HMI tags "Default tag table"
   "buttonView" : Bool, internal
   "messageView" : Bool, internal
   "RPA30R_LCDSwitchAutomat_Manual" : Bool = PLC "RPA30R_LCDSwitchAutomat_Manual", 100 ms
   "RPA30R_light" : Bool = PLC "RPA30R_light", 100 ms
   "RPA30_DataBlock_RPA30_Start" : Bool, 100 ms
   "RPA30_DataBlock_RPA30_scannedFrameBareCode" : String[254], 100 ms
   "RPA30_DataBlock_RPA30_cyclusState" : UInt, 100 ms
   "RPA30_DataBlock_RPA30_scannedData" : String[254], 100 ms
   "outputStatePageChose" : Int, internal
   "ipnut_page_switch" : Int, internal
   "inputStatePageChose" : Int, internal
   "RPA30R_RoofRotationSensorYL" : Bool = PLC "RPA30R_RoofRotationSensorYL", 100 ms
   "RPA30R_RoofRotationSensorYAtOperator" : Bool = PLC "RPA30R_RoofRotationSensorYAtOperator", 100 ms
   "RPA30R_RoofRotationSensorYR" : Bool = PLC "RPA30R_RoofRotationSensorYR", 100 ms
   "RPA30R_RoofRotationSensorYFromOperator" : Bool = PLC "RPA30R_RoofRotationSensorYFromOperator", 100 ms
   "RPA30R_PositionCylinderSensorUnlockY" : Bool = PLC "RPA30R_PositionCylinderSensorUnlockY", 100 ms
   "RPA30R_PositionCylinderSensorLockY" : Bool = PLC "RPA30R_PositionCylinderSensorLockY", 100 ms
   "RPA30R_SensorIFMLeftTriggerOut" : Bool = PLC "RPA30R_SensorIFMLeftTriggerOut", 100 ms
   "RPA30R_SensorIFMLeftReadyOut" : Bool = PLC "RPA30R_SensorIFMLeftReadyOut", 100 ms
   "RPA30R_SensorIFMLeftOut" : Bool = PLC "RPA30R_SensorIFMLeftOut", 100 ms
   "RPA30R_SensorIFMRightTriggerOut" : Bool = PLC "RPA30R_SensorIFMRightTriggerOut", 100 ms
   "RPA30R_SensorIFMRightReadyOut" : Bool = PLC "RPA30R_SensorIFMRightReadyOut", 100 ms
   "RPA30R_SensorIFMRightOut" : Bool = PLC "RPA30R_SensorIFMRightOut", 100 ms
   "RPA30R_ValveCylinderYLock" : Bool = PLC "RPA30R_ValveCylinderYLock", 100 ms
   "RPA30R_SensorIFMLeftTrigger" : Bool = PLC "RPA30R_SensorIFMLeftTrigger", 100 ms
   "RPA30R_SensorIFMLeft_Input_1" : Bool = PLC "RPA30R_SensorIFMLeft_Input_1", 100 ms
   "RPA30R_SensorIFMLeft_Input_2" : Bool = PLC "RPA30R_SensorIFMLeft_Input_2", 100 ms
   "RPA30R_SensorIFMRightTrigger" : Bool = PLC "RPA30R_SensorIFMRightTrigger", 100 ms
   "RPA30R_SensorIFMRight_Input_1" : Bool = PLC "RPA30R_SensorIFMRight_Input_1", 100 ms
   "RPA30R_SensorIFMRight_Input_2" : Bool = PLC "RPA30R_SensorIFMRight_Input_2", 100 ms
   "RPA30R_PrimerPA10SensorPadLeft" : Bool = PLC "RPA30R_PrimerPA10SensorPadLeft", 100 ms
   "RPA30R_PrimerPA10SensorPadRight" : Bool = PLC "RPA30R_PrimerPA10SensorPadRight", 100 ms
   "RPA30R_PrimerPA10SensorFelt" : Bool = PLC "RPA30R_PrimerPA10SensorFelt", 100 ms
   "RPA30R_PrimerPA30SensorRemover208" : Bool = PLC "RPA30R_PrimerPA30SensorRemover208", 100 ms
   "RPA30R_PrimerPA30SensorFeltEmpty" : Bool = PLC "RPA30R_PrimerPA30SensorFeltEmpty", 100 ms
   "RPA30R_LCDButtonStart" : Bool = PLC "RPA30R_LCDButtonStart", 100 ms
   "RPA30R_LCDButtonConfirmSignal" : Bool = PLC "RPA30R_LCDButtonConfirmSignal", 100 ms
   "RPA30R_PrimerPA30SensorBottleRemover208" : Bool = PLC "RPA30R_PrimerPA30SensorBottleRemover208", 100 ms
   "RPA30R_PrimerPA30SensorBottlePrimer207" : Bool = PLC "RPA30R_PrimerPA30SensorBottlePrimer207", 100 ms
   "RPA30R_Beacon_1_LCDPanelGreen" : Bool = PLC "RPA30R_Beacon_1_LCDPanelGreen", 100 ms
   "RPA30R_Beacon_1_LCDPanelOrange" : Bool = PLC "RPA30R_Beacon_1_LCDPanelOrange", 100 ms
   "RPA30R_Beacon_1_LCDPanelRed" : Bool = PLC "RPA30R_Beacon_1_LCDPanelRed", 100 ms
   "RPA30R_Beacon_1_LCDPanelSiren" : Bool = PLC "RPA30R_Beacon_1_LCDPanelSiren", 100 ms
   "RPA30R_Beacon_2_PrimerBoxGreen" : Bool = PLC "RPA30R_Beacon_2_PrimerBoxGreen", 100 ms
   "RPA30R_Beacon_2_PrimerBoxOrange" : Bool = PLC "RPA30R_Beacon_2_PrimerBoxOrange", 100 ms
   "RPA30R_Beacon_2_PrimerBoxRed" : Bool = PLC "RPA30R_Beacon_2_PrimerBoxRed", 100 ms
   "RPA30R_Beacon_2_PrimerBoxSiren" : Bool = PLC "RPA30R_Beacon_2_PrimerBoxSiren", 100 ms
   "RPA30R_PrimerPA30GreenReady" : Bool = PLC "RPA30R_PrimerPA30GreenReady", 100 ms
   "RPA30R_PrimerPA30GreenFelt" : Bool = PLC "RPA30R_PrimerPA30GreenFelt", 100 ms
   "RPA30R_PrimerPA30GreenRemover208" : Bool = PLC "RPA30R_PrimerPA30GreenRemover208", 100 ms
   "RPA30R_PrimerPA30GreenPrimer207" : Bool = PLC "RPA30R_PrimerPA30GreenPrimer207", 100 ms
   "RPA30R_PrimerPA30RedNotReady" : Bool = PLC "RPA30R_PrimerPA30RedNotReady", 100 ms
   "RPA30R_PrimerPA30RedChangePad" : Bool = PLC "RPA30R_PrimerPA30RedChangePad", 100 ms
   "RPA30R_LEDGreenSart" : Bool = PLC "RPA30R_LEDGreenSart", 100 ms
   "RPA30R_LedBlueConfirm" : Bool = PLC "RPA30R_LedBlueConfirm", 100 ms
   "RPA30_DataBlock_RPA30_failStateLock" : Int, 100 ms
   "Clock_0.5Hz" : Bool = PLC "Clock_0.5Hz", 100 ms
   "RPA30_DataBlock_RPA30_bigFailStateLock" : Int, 100 ms
   "RPA30_DataBlock_RPA30_ErrorStateLock" : Int, 100 ms
   "RPA30_DataBlock_RPA30_fatalErrorStateLock" : Int, 100 ms
   "RPA30_IFM_point_checking_DB_points" : Int, 100 ms
   "manual_output_page_switch" : Int, internal
   "input_output_switch" : Bool, internal
   "output_page_switch" : Int, internal
   "PLC_datablock_stations_configuration" : Byte, 1 s
   "configuration_choose" : Int, internal
   "RPA30_DataBlock_RPA30_show_points_hmi" : Byte, 100 ms
   "RPA30_DataBlock_RPA30_actual_instruction_index" : Byte, 1 s
   "RPA30_DataBlock_RPA30_show_smile" : Bool, 100 ms
   "RPA30_DataBlock_RPA30_show_pad_left" : Bool, 100 ms
   "RPA30_DataBlock_RPA30_show_pad_right" : Bool, 100 ms
   "RPA30_DataBlock_pa30_bottle_cyclus_replace" : UInt, 1 s
   "RPA30_DataBlock_pa30_bottle_timing" : LInt, 1 s
   "RPA30_DataBlock_pa30_keyence_switch" : Bool, 1 s

text list "RPA30_InstructionList": 0 ''; 1 ''; 4 ''; 5 ''; 6 ''; 7 ''; 9 ''; 16 ''; 17 ''; 18 ''; 19 ''; 20 ''; 21 ''; 22 ''; 23 ''; 24 ''; 25 ''; 26 ''; 27 ''; 28 ''

text list "pa30_fail_list": 200 ''; 210 ''; 100 ''; 300 ''

text list "PA30_error_list": 1000 ''; 25000 ''; 26000 ''; 24000 ''; 23000 ''; 22000 ''; 400 ''; 401 ''; 402 ''; 403 ''; 155 ''

text list "PA30_fatal_error_list": 150 ''; 160 ''; 190 ''

text list "RPA30_station_configuration": 0 ''; 1 ''; 2 ''

screen "Home" 800x480
   TextField "Text field_3" at 325,5 size 300x40
   TextField "Text field_2" at 2,85 size 70x40
   TextField "Text field_4" at 73,85 size 70x40
   TextField "Text field_5" at 335,130 size 130x25
   TextField "Text field_6" at 20,171 size 330x22
   TextField "Text field_7" at 20,201 size 330x22
   TextField "Text field_8" at 20,231 size 330x22
   TextField "Text field_9" at 20,261 size 330x22
   TextField "Text field_10" at 20,291 size 330x22
   TextField "Text field_11" at 20,321 size 330x22
   TextField "Text field_12" at 20,351 size 330x22
   TextField "Text field_13" at 20,381 size 330x22
   TextField "Text field_14" at 410,171 size 330x22
   TextField "Text field_15" at 410,201 size 330x22
   TextField "Text field_16" at 410,231 size 330x22
   TextField "Text field_17" at 410,261 size 330x22
   TextField "Text field_18" at 410,291 size 330x22
   TextField "Text field_19" at 410,321 size 330x22
   TextField "Text field_20" at 410,351 size 330x22
   TextField "Text field_21" at 410,381 size 330x22
   Button "Button_1" at 640,420 size 80x60
   Button "HmiScreenItemData_1" at 0,420 size 80x60
   Button "HmiScreenItemData_2" at 400,420 size 80x60
   Button "Button_2" at 560,420 size 80x60
   Button "Button_6" at 720,420 size 80x60
   DateTimeField "Date/time field_1" at 650,27 size 150x25
   DateTimeField "Date/time field_2" at 650,0 size 150x28
   TextField "Text field_1" at 0,0 size 300x50
   Button "HmiScreenItemData_3" at 240,420 size 80x60
   Button "HmiScreenItemData_4" at 320,420 size 80x60
   Button "Button_3" at 480,420 size 80x60
   Button "HmiScreenItemData_5" at 80,420 size 80x60
   Button "HmiScreenItemData_6" at 160,420 size 80x60
   Button "Button_11" at 0,420 size 80x60
   Button "Button_12" at 80,420 size 80x60
   Button "Button_13" at 160,420 size 80x60
   Button "Button_14" at 240,420 size 80x60
   Button "Button_15" at 320,420 size 80x60
   Button "Button_16" at 400,420 size 80x60
   Button "Button_17" at 480,420 size 80x60
   Button "Button_18" at 560,420 size 80x60
   Button "Button_19" at 640,420 size 80x60
   Button "Button_20" at 720,420 size 80x60
   TextField "Text field_22" at 64,67 size 129x22
   AlarmView "Alarm view_1" at 60,90 size 680x320
   Button "Button_9" at 715,65 size 25x25
   TextField "Text field_37" at 360,54 size 120x25

screen "I0-State" 800x480
   TextField "Text field_3" at 325,5 size 300x40
   Button "Button_1" at 640,420 size 80x60
   Button "Button_4" at 160,420 size 80x60
   Button "HmiScreenItemData_3" at 400,420 size 80x60
   Button "Button_2" at 560,420 size 80x60
   Button "Button_6" at 720,420 size 80x60
   Button "HmiScreenItemData_2" at 240,420 size 80x60
   Button "HmiScreenItemData_4" at 320,420 size 80x60
   TextField "Text field_1" at 0,0 size 300x50
   DateTimeField "Date/time field_2" at 650,0 size 150x28
   DateTimeField "Date/time field_1" at 650,27 size 150x25
   Button "HmiScreenItemData_1" at 0,420 size 80x60
   Button "Button_3" at 480,420 size 80x60
   Button "Button_5" at 80,420 size 80x60
   Button "input_back" at 20,52 size 90x25
   Button "input_next" at 690,52 size 90x25
   Button "output_back" at 20,52 size 90x25
   Button "output_next" at 690,52 size 90x25
   TextField "Text field_2" at 20,85 size 330x22
   TextField "Text field_4" at 20,115 size 330x22
   TextField "Text field_5" at 20,145 size 330x22
   TextField "Text field_6" at 20,175 size 330x22
   TextField "Text field_7" at 20,205 size 330x22
   TextField "Text field_8" at 20,235 size 330x22
   TextField "Text field_9" at 20,265 size 330x22
   TextField "Text field_10" at 20,295 size 330x22
   TextField "Text field_11" at 20,325 size 330x22
   TextField "Text field_12" at 20,355 size 330x22
   TextField "Text field_13" at 20,385 size 330x22
   TextField "Text field_14" at 410,85 size 330x22
   TextField "Text field_15" at 410,115 size 330x22
   TextField "Text field_16" at 410,145 size 330x22
   TextField "Text field_17" at 410,175 size 330x22
   TextField "Text field_18" at 410,205 size 330x22
   TextField "Text field_19" at 410,235 size 330x22
   TextField "Text field_20" at 410,265 size 330x22
   TextField "Text field_21" at 410,295 size 330x22
   TextField "Text field_22" at 410,325 size 330x22
   TextField "Text field_23" at 410,355 size 330x22
   TextField "Text field_24" at 410,385 size 330x22
   Button "Button_11" at 0,420 size 80x60
   Button "Button_12" at 80,420 size 80x60
   Button "Button_13" at 160,420 size 80x60
   Button "Button_14" at 240,420 size 80x60
   Button "Button_15" at 320,420 size 80x60
   Button "Button_16" at 400,420 size 80x60
   Button "Button_17" at 480,420 size 80x60
   Button "Button_18" at 560,420 size 80x60
   Button "Button_19" at 640,420 size 80x60
   Button "Button_20" at 720,420 size 80x60
   TextField "Text field_25" at 64,67 size 129x22
   AlarmView "Alarm view_1" at 60,90 size 680x320
   Button "Button_9" at 715,65 size 25x25
   TextField "Text field_26" at 20,85 size 330x22
   TextField "Text field_27" at 20,115 size 330x22
   TextField "Text field_28" at 20,145 size 330x22
   TextField "Text field_29" at 20,175 size 330x22
   TextField "Text field_30" at 20,205 size 330x22
   TextField "Text field_31" at 20,235 size 330x22
   TextField "Text field_32" at 20,265 size 330x22
   TextField "Text field_33" at 20,295 size 330x22
   TextField "Text field_34" at 20,325 size 330x22
   TextField "Text field_35" at 20,355 size 330x22
   TextField "Text field_36" at 20,385 size 330x22
   TextField "Text field_37" at 410,85 size 330x22
   TextField "Text field_38" at 410,115 size 330x22
   TextField "Text field_39" at 410,145 size 330x22
   TextField "Text field_40" at 410,175 size 330x22
   TextField "Text field_41" at 410,205 size 330x22
   TextField "Text field_42" at 410,235 size 330x22
   TextField "Text field_43" at 410,265 size 330x22
   TextField "Text field_44" at 410,295 size 330x22
   TextField "Text field_45" at 410,325 size 330x22
   TextField "Text field_46" at 410,355 size 330x22
   TextField "Text field_47" at 410,385 size 330x22
   TextField "Text field_48" at 20,85 size 330x22
   TextField "Text field_49" at 20,85 size 330x22
   TextField "Text field_50" at 360,54 size 120x25

screen "Main_page" 800x480
   Button "HmiScreenItemData_1" at 80,420 size 80x60
   TextField "Text field_2" at 0,85 size 800x25
   TextField "Text field_3" at 325,5 size 300x40
   Button "Button_4" at 480,420 size 80x60
   Button "Button_5" at 640,420 size 80x60
   Button "Button_1" at 0,420 size 80x60
   Button "Button_7" at 400,420 size 80x60
   Button "HmiScreenItemData_2" at 160,420 size 80x60
   Button "Button_3" at 560,420 size 80x60
   Button "Button_6" at 720,420 size 80x60
   Button "HmiScreenItemData_3" at 240,420 size 80x60
   Button "HmiScreenItemData_4" at 320,420 size 80x60
   TextField "Text field_1" at 0,0 size 300x50
   DateTimeField "Date/time field_2" at 650,0 size 150x28
   DateTimeField "Date/time field_1" at 650,27 size 150x25
   SymbolicIOField "Symbolic I/O field_1" at 10,110 size 780x90
   Button "HmiScreenItemData_5" at 80,420 size 80x60
   SymbolicIOField "Symbolic I/O field_6" at 171,50 size 169x32
   TextField "Text field_56" at 11,51 size 143x27
   Button "Button_2" at 400,420 size 80x60
   Button "Button_11" at 0,420 size 80x60
   Button "Button_12" at 80,420 size 80x60
   Button "Button_13" at 160,420 size 80x60
   Button "Button_14" at 240,420 size 80x60
   Button "Button_15" at 320,420 size 80x60
   Button "Button_16" at 400,420 size 80x60
   Button "Button_17" at 480,420 size 80x60
   Button "Button_18" at 560,420 size 80x60
   Button "Button_19" at 640,420 size 80x60
   Button "Button_20" at 720,420 size 80x60
   GraphicView "Graphic view_1" at 320,228 size 180x180
   TextField "Text field_5" at 64,67 size 129x22
   AlarmView "Alarm view_1" at 60,90 size 680x320
   Button "Button_9" at 715,65 size 25x25
   SymbolicIOField "Symbolic I/O field_2" at 0,170 size 800x110
   SymbolicIOField "Symbolic I/O field_3" at 0,170 size 800x110
   SymbolicIOField "Symbolic I/O field_4" at 0,170 size 800x110
   SymbolicIOField "Symbolic I/O field_5" at 0,170 size 800x110
   TextField "Text field_10" at 165,322 size 22x37
   TextField "Text field_11" at 279,323 size 22x37
   TextField "Text field_12" at 392,323 size 22x37
   TextField "Text field_13" at 494,322 size 22x37
   TextField "Text field_14" at 613,323 size 22x37
   TextField "Text field_6" at 163,255 size 22x37
   TextField "Text field_7" at 392,255 size 22x37
   TextField "Text field_8" at 613,255 size 22x37
   TextField "Text field_37" at 360,54 size 120x25
   GraphicView "Graphic view_2" at 207,225 size 345x187
   GraphicView "Graphic view_3" at 260,225 size 345x187
   TextField "Text field_4" at 299,290 size 237x43

screen "Scanner" 800x480
   TextField "Text field_3" at 325,5 size 300x40
   IOField "I/O field_1" at 10,118 size 780x32
   TextField "Text field_2" at 10,86 size 141x22
   Button "Button_1" at 640,420 size 80x60
   Button "HmiScreenItemData_3" at 400,420 size 80x60
   Button "Button_2" at 560,420 size 80x60
   Button "Button_6" at 720,420 size 80x60
   DateTimeField "Date/time field_2" at 650,0 size 150x28
   TextField "Text field_1" at 0,0 size 300x50
   DateTimeField "Date/time field_1" at 650,27 size 150x25
   Button "HmiScreenItemData_2" at 240,420 size 80x60
   Button "HmiScreenItemData_4" at 320,420 size 80x60
   Button "HmiScreenItemData_1" at 0,420 size 80x60
   Button "HmiScreenItemData_5" at 480,420 size 80x60
   Button "HmiScreenItemData_6" at 160,420 size 80x60
   Button "HmiScreenItemData_7" at 80,420 size 80x60
   Button "Button_3" at 27,167 size 96x32
   Button "Button_11" at 0,420 size 80x60
   Button "Button_12" at 80,420 size 80x60
   Button "Button_13" at 160,420 size 80x60
   Button "Button_14" at 240,420 size 80x60
   Button "Button_15" at 320,420 size 80x60
   Button "Button_16" at 400,420 size 80x60
   Button "Button_17" at 480,420 size 80x60
   Button "Button_18" at 560,420 size 80x60
   Button "Button_19" at 640,420 size 80x60
   Button "Button_20" at 720,420 size 80x60
   TextField "Text field_5" at 64,67 size 129x22
   AlarmView "Alarm view_1" at 60,90 size 680x320
   Button "Button_9" at 715,65 size 25x25
   TextField "Text field_37" at 360,54 size 120x25

screen "Manual" 800x480
   TextField "Text field_3" at 325,5 size 300x40
   Button "Button_4" at 18,85 size 50x50
   Button "Button_12" at 730,85 size 50x50
   Button "Button_1" at 640,420 size 80x60
   Button "HmiScreenItemData_1" at 0,420 size 80x60
   Button "Button_6" at 720,420 size 80x60
   Button "Button_34" at 400,420 size 80x60
   Button "HmiScreenItemData_3" at 240,420 size 80x60
   Button "HmiScreenItemData_4" at 320,420 size 80x60
   TextField "Text field_1" at 0,0 size 300x50
   DateTimeField "Date/time field_2" at 650,0 size 150x28
   DateTimeField "Date/time field_1" at 650,27 size 150x25
   Button "Button_5" at 160,420 size 80x60
   Button "Button_3" at 480,420 size 80x60
   Button "Button_7" at 80,420 size 80x60
   Button "Button_2" at 560,420 size 80x60
   Button "Button_23" at 0,420 size 80x60
   Button "Button_24" at 80,420 size 80x60
   Button "Button_25" at 160,420 size 80x60
   Button "Button_26" at 240,420 size 80x60
   Button "Button_27" at 320,420 size 80x60
   Button "Button_28" at 400,420 size 80x60
   Button "Button_29" at 480,420 size 80x60
   Button "Button_30" at 560,420 size 80x60
   Button "Button_31" at 640,420 size 80x60
   Button "Button_32" at 720,420 size 80x60
   TextField "Text field_8" at 64,67 size 129x22
   AlarmView "Alarm view_1" at 60,90 size 680x320
   Button "Button_33" at 715,65 size 25x25
   Switch "Switch_15" at 717,149 size 64x32
   Switch "Switch_16" at 717,185 size 64x32
   Switch "Switch_17" at 717,221 size 64x32
   Switch "Switch_18" at 717,257 size 64x32
   Switch "Switch_19" at 717,293 size 64x32
   Switch "Switch_20" at 718,328 size 64x32
   Switch "Switch_21" at 719,364 size 64x32
   TextField "Text field_22" at 493,149 size 200x32
   TextField "Text field_23" at 493,181 size 200x32
   TextField "Text field_24" at 492,221 size 200x32
   TextField "Text field_25" at 493,289 size 200x32
   TextField "Text field_26" at 493,257 size 200x32
   TextField "Text field_27" at 493,328 size 200x32
   TextField "Text field_28" at 493,360 size 200x32
   Switch "Switch_22" at 300,149 size 64x32
   Switch "Switch_23" at 300,185 size 64x32
   Switch "Switch_24" at 300,221 size 64x32
   Switch "Switch_25" at 300,257 size 64x32
   Switch "Switch_26" at 300,293 size 64x32
   Switch "Switch_27" at 301,328 size 64x32
   Switch "Switch_28" at 302,364 size 64x32
   TextField "Text field_29" at 76,149 size 200x32
   TextField "Text field_30" at 76,181 size 200x32
   TextField "Text field_31" at 75,221 size 200x32
   TextField "Text field_32" at 76,289 size 200x32
   TextField "Text field_33" at 76,257 size 200x32
   TextField "Text field_34" at 76,328 size 200x32
   TextField "Text field_35" at 76,360 size 200x32
   Switch "Switch_1" at 717,149 size 64x32
   Switch "Switch_2" at 717,185 size 64x32
   TextField "Text field_7" at 493,149 size 200x32
   TextField "Text field_9" at 493,181 size 200x32
   Switch "Switch_8" at 300,149 size 64x32
   Switch "Switch_9" at 300,185 size 64x32
   Switch "Switch_10" at 300,221 size 64x32
   Switch "Switch_11" at 300,257 size 64x32
   Switch "Switch_12" at 300,293 size 64x32
   Switch "Switch_13" at 301,328 size 64x32
   Switch "Switch_14" at 302,364 size 64x32
   TextField "Text field_15" at 76,149 size 200x32
   TextField "Text field_16" at 76,181 size 200x32
   TextField "Text field_17" at 75,221 size 200x32
   TextField "Text field_18" at 37,289 size 239x32
   TextField "Text field_19" at 26,257 size 250x32
   TextField "Text field_20" at 29,328 size 247x32
   TextField "Text field_21" at 44,360 size 232x32
   TextField "Text field_37" at 360,54 size 120x25

screen "System" 800x480
   TextField "Text field_3" at 325,5 size 300x40
   TextField "Text field_2" at 300,86 size 200x27
   Button "Button_4" at 10,290 size 170x60
   Button "Button_5" at 10,355 size 170x60
   Button "Button_7" at 213,290 size 170x60
   Button "Button_8" at 416,290 size 170x60
   Button "Button_9" at 620,290 size 170x60
   Button "Button_11" at 213,355 size 170x60
   Button "Button_12" at 416,355 size 170x60
   Button "Button_13" at 620,355 size 170x60
   AlarmView "Alarm view_1" at 10,115 size 780x170
   Button "HmiScreenItemData_1" at 0,420 size 80x60
   Button "Button_3" at 160,420 size 80x60
   Button "Button_14" at 240,420 size 80x60
   Button "Button_15" at 320,420 size 80x60
   Button "Button_16" at 400,420 size 80x60
   Button "Button_2" at 560,420 size 80x60
   Button "Button_1" at 640,420 size 80x60
   Button "Button_6" at 720,420 size 80x60
   TextField "Text field_1" at 0,0 size 300x50
   DateTimeField "Date/time field_2" at 650,0 size 150x28
   DateTimeField "Date/time field_1" at 650,27 size 150x25
   Button "Button_10" at 80,420 size 80x60
   Button "Button_17" at 480,420 size 80x60
   TextField "Text field_37" at 360,54 size 120x25

screen "Station_configuration" 800x480
   TextField "Text field_3" at 325,5 size 300x40
   Button "Button_1" at 640,420 size 80x60
   Button "HmiScreenItemData_1" at 0,420 size 80x60
   Button "Button_6" at 720,420 size 80x60
   Button "Button_34" at 400,420 size 80x60
   Button "HmiScreenItemData_4" at 320,420 size 80x60
   TextField "Text field_1" at 0,0 size 300x50
   DateTimeField "Date/time field_2" at 650,0 size 150x28
   DateTimeField "Date/time field_1" at 650,27 size 150x25
   Button "Button_5" at 160,420 size 80x60
   Button "Button_3" at 480,420 size 80x60
   Button "Button_7" at 80,420 size 80x60
   Button "Button_2" at 560,420 size 80x60
   SymbolicIOField "Symbolic I/O field_1" at 33,194 size 310x65
   TextField "Text field_2" at 33,159 size 192x27
   Button "Button_4" at 355,195 size 90x65
   SymbolicIOField "Symbolic I/O field_2" at 457,195 size 310x65
   TextField "Text field_4" at 457,159 size 225x27
   Switch "Switch_1" at 370,326 size 64x32
   TextField "Text field_5" at 222,288 size 223x23
   Button "HmiScreenItemData_2" at 240,420 size 80x60
   TextField "Text field_37" at 360,54 size 120x25

screen "chemical_setup" 800x480
   Button "HmiScreenItemData_3" at 400,420 size 80x60
   Button "Button_2" at 560,420 size 80x60
   Button "Button_6" at 720,420 size 80x60
   DateTimeField "Date/time field_2" at 650,0 size 150x28
   TextField "Text field_1" at 0,0 size 300x50
   DateTimeField "Date/time field_1" at 650,27 size 150x25
   Button "HmiScreenItemData_2" at 240,420 size 80x60
   Button "HmiScreenItemData_4" at 320,420 size 80x60
   Button "HmiScreenItemData_1" at 0,420 size 80x60
   Button "HmiScreenItemData_5" at 480,420 size 80x60
   Button "HmiScreenItemData_6" at 160,420 size 80x60
   Button "HmiScreenItemData_7" at 80,420 size 80x60
   IOField "I/O field_1" at 87,130 size 341x44
   IOField "I/O field_2" at 87,237 size 338x44
   TextField "Text field_2" at 85,100 size 137x25
   TextField "Text field_3" at 87,206 size 111x25
   TextField "Text field_4" at 435,245 size 93x20
   Button "Button_1" at 640,420 size 80x60
   Button "Button_11" at 0,420 size 80x60
   Button "Button_12" at 80,420 size 80x60
   Button "Button_13" at 160,420 size 80x60
   Button "Button_14" at 240,420 size 80x60
   Button "Button_15" at 320,420 size 80x60
   Button "Button_16" at 400,420 size 80x60
   Button "Button_17" at 480,420 size 80x60
   Button "Button_18" at 560,420 size 80x60
   Button "Button_19" at 640,420 size 80x60
   Button "Button_20" at 720,420 size 80x60
   TextField "Text field_5" at 64,67 size 129x22
   Button "Button_9" at 715,65 size 25x25
   AlarmView "Alarm view_1" at 60,90 size 680x320
   TextField "Text field_37" at 360,54 size 120x25

screen "User_management" 800x480
   TextField "Text field_3" at 325,5 size 300x40
   Button "HmiScreenItemData_1" at 0,420 size 80x60
   Button "Button_3" at 160,420 size 80x60
   Button "Button_14" at 240,420 size 80x60
   Button "Button_15" at 320,420 size 80x60
   Button "Button_16" at 400,420 size 80x60
   Button "Button_17" at 480,420 size 80x60
   Button "Button_2" at 560,420 size 80x60
   Button "Button_1" at 640,420 size 80x60
   TextField "Text field_1" at 0,0 size 300x50
   DateTimeField "Date/time field_2" at 650,0 size 150x28
   DateTimeField "Date/time field_1" at 650,27 size 150x25
   Button "Button_10" at 80,420 size 80x60
   UserView "User view_1" at 20,92 size 758x304
   Button "Button_4" at 720,420 size 80x60
   TextField "Text field_37" at 360,54 size 120x25
*)

(* ===== HMI "HMI_RT_4" =====
connection "HMI_Connection_4": ETHERNET, SMART_S7_1500_OMS

HMI tags "Default tag table"
   "buttonView" : Bool, internal
   "messageView" : Bool, internal
   "RPA60R_LCDSwitchAutomat_Manual" : Bool = PLC "RPA60R_LCDSwitchAutomat_Manual", 100 ms
   "RPA60R_light" : Bool = PLC "RPA60R_light", 100 ms
   "RPA60_DataBlock_RPA60_Start" : Bool, 100 ms
   "RPA60_DataBlock_RPA60_cyclusState" : UInt, 100 ms
   "RPA60_DataBlock_RPA60_scannedFrameBareCode" : String[254], 100 ms
   "RPA60_DataBlock_RPA60_failStateLock" : Int, 100 ms
   "RPA60_DataBlock_RPA60_scanedData" : String[254], 100 ms
   "inputOutputStatePageChose" : Int, internal
   "RPA60R_RoofRotationSensorYL" : Bool = PLC "RPA60R_RoofRotationSensorYL", 100 ms
   "RPA60R_RoofRotationSensorYAtOperator" : Bool = PLC "RPA60R_RoofRotationSensorYAtOperator", 100 ms
   "RPA60R_RoofRotationSensorYR" : Bool = PLC "RPA60R_RoofRotationSensorYR", 100 ms
   "RPA60R_RoofRotationSensorYFromOperator" : Bool = PLC "RPA60R_RoofRotationSensorYFromOperator", 100 ms
   "RPA60R_valvePositionSensorUnlockY" : Bool = PLC "RPA60R_valvePositionSensorUnlockY", 100 ms
   "RPA60R_valvePositionSensorLockY" : Bool = PLC "RPA60R_valvePositionSensorLockY", 100 ms
   "RPA60R_SenzorLoaderPresenceLeft581" : Bool = PLC "RPA60R_SenzorLoaderPresenceLeft581", 100 ms
   "RPA60R_SenzorLoaderPresenceRight581" : Bool = PLC "RPA60R_SenzorLoaderPresenceRight581", 100 ms
   "RPA60R_SenzorLoaderPresenceLeft582" : Bool = PLC "RPA60R_SenzorLoaderPresenceLeft582", 100 ms
   "RPA60R_SenzorLoaderPresenceRear582" : Bool = PLC "RPA60R_SenzorLoaderPresenceRear582", 100 ms
   "RPA60R_SenzorLoaderPresenceRight582" : Bool = PLC "RPA60R_SenzorLoaderPresenceRight582", 100 ms
   "RPA60R_SenzorSealPresenceLeft581" : Bool = PLC "RPA60R_SenzorSealPresenceLeft581", 100 ms
   "RPA60R_SenzorSealPresenceRear581" : Bool = PLC "RPA60R_SenzorSealPresenceRear581", 100 ms
   "RPA60R_SenzorSealPresenceRight581" : Bool = PLC "RPA60R_SenzorSealPresenceRight581", 100 ms
   "RPA60R_SenzorSealPresenceLeft582" : Bool = PLC "RPA60R_SenzorSealPresenceLeft582", 100 ms
   "RPA60R_SenzorSealPresenceRear582" : Bool = PLC "RPA60R_SenzorSealPresenceRear582", 100 ms
   "RPA60R_SenzorSealPresenceRight582" : Bool = PLC "RPA60R_SenzorSealPresenceRight582", 100 ms
   "RPA60R_SenzorVacuum" : Bool = PLC "RPA60R_SenzorVacuum", 100 ms
   "RPA60R_ValveCylinderYLock" : Bool = PLC "RPA60R_ValveCylinderYLock", 100 ms
   "RPA60R_LCDButtonStart" : Bool = PLC "RPA60R_LCDButtonStart", 100 ms
   "RPA60R_LCDButtonConfirmSignal" : Bool = PLC "RPA60R_LCDButtonConfirmSignal", 100 ms
   "RPA60R_Beacon_1_LCDPanelGreen" : Bool = PLC "RPA60R_Beacon_1_LCDPanelGreen", 100 ms
   "RPA60R_Beacon_1_LCDPanelOrange" : Bool = PLC "RPA60R_Beacon_1_LCDPanelOrange", 100 ms
   "RPA60R_Beacon_1_LCDPanelRed" : Bool = PLC "RPA60R_Beacon_1_LCDPanelRed", 100 ms
   "RPA60R_Beacon_1_LCDPanelSiren" : Bool = PLC "RPA60R_Beacon_1_LCDPanelSiren", 100 ms
   "RPA60R_LEDGreenSart" : Bool = PLC "RPA60R_LEDGreenSart", 100 ms
   "RPA60R_LedBlueConfirm" : Bool = PLC "RPA60R_LedBlueConfirm", 100 ms
   "RPA60R_VacuumSwitch" : Bool = PLC "RPA60R_VacuumSwitch", 100 ms
   "RPA60R_LEDRoller" : Bool = PLC "RPA60R_LEDRoller", 100 ms
   "RPA60R_SenzorRoller" : Bool = PLC "RPA60R_SenzorRoller", 100 ms
   "RPA30R_Beacon_1_LCDPanelSiren" : Bool = PLC "RPA30R_Beacon_1_LCDPanelSiren", 100 ms
   "RPA60_DataBlock_RPA60_bigFailStateLock" : Int, 1 s
   "RPA60_DataBlock_RPA60_fatalErrorStateLock" : Int, 1 s
   "RPA60_DataBlock_RPA60_ErrorStateLock" : Int, 1 s
   "Clock_0.5Hz" : Bool = PLC "Clock_0.5Hz", 1 s
   "RPA60_DataBlock_RPA60_printEnable" : Bool, 1 s
   "input_output_switch" : Bool, internal
   "output_switch_page" : Int, internal
   "input_switch_page" : Int, internal
   "PLC_datablock_stations_configuration" : Byte, 1 s
   "RPA60_DataBlock_RPA60_hmi_instruction_index" : Byte, 1 s
   "RPA60_DataBlock_RPA60_show_smile" : Bool, 1 s
   "RPA60_DataBlock_RPA60_number_of_check" : Byte, 1 s
   "RPA60_DataBlock_RPA60_show_check_button" : Bool, 1 s
   "RPA60_DataBlock_RPA60_station_configuration" : Byte, 1 s
   "choose_configuration" : Int, internal
   "RPA60_DataBlock_RPA60_hardware_configuration" : Byte, 1 s
   "DB_RPA60_CAM_RPA60_ENABLE_CAMERAS" : Bool, 500 ms

text list "PA60_instructionList": 0 ''; 3 ''; 7 ''; 8 ''; 9 ''; 24 ''; 26 ''; 27 ''; 23 ''; 28 ''; 11 ''; 29 ''; 30 ''; 39 ''; 40 ''; 41 ''

text list "PA60_error_list": 1000 ''; 26000 ''; 25000 ''; 24000 ''; 23000 ''; 20000 ''; 21000 ''; 27000 ''

text list "PA60_fatal_error_list": 170 ''; 150 ''; 180 ''; 230 ''; 293 ''; 294 ''; 190 ''

text list "PA60_big_fail_list": 120 ''

text list "RPA60_station_configuration": 0 ''; 1 ''; 2 ''

text list "RPA60_hardware_configuration": 0 ''; 1 ''; 3..255 ''; 2 ''

screen "Home" 800x480
   TextField "Text field_3" at 325,5 size 300x40
   TextField "Text field_2" at 2,85 size 70x40
   TextField "Text field_5" at 335,130 size 130x25
   TextField "Text field_6" at 20,171 size 330x22
   TextField "Text field_7" at 20,201 size 330x22
   Button "Button_1" at 640,420 size 80x60
   Button "HmiScreenItemData_1" at 0,420 size 80x60
   Button "HmiScreenItemData_2" at 400,420 size 80x60
   Button "Button_2" at 560,420 size 80x60
   Button "Button_6" at 720,420 size 80x60
   DateTimeField "Date/time field_1" at 650,27 size 150x25
   DateTimeField "Date/time field_2" at 650,0 size 150x28
   TextField "Text field_1" at 0,0 size 300x50
   Button "HmiScreenItemData_3" at 240,420 size 80x60
   Button "HmiScreenItemData_4" at 320,420 size 80x60
   Button "Button_3" at 480,420 size 80x60
   Button "HmiScreenItemData_5" at 80,420 size 80x60
   Button "HmiScreenItemData_6" at 160,420 size 80x60
   IOField "I/O field_1" at 73,85 size 70x40
   Button "Button_11" at 0,420 size 80x60
   Button "Button_12" at 80,420 size 80x60
   Button "Button_13" at 160,420 size 80x60
   Button "Button_14" at 240,420 size 80x60
   Button "Button_15" at 320,420 size 80x60
   Button "Button_16" at 400,420 size 80x60
   Button "Button_17" at 480,420 size 80x60
   Button "Button_18" at 560,420 size 80x60
   Button "Button_19" at 640,420 size 80x60
   Button "Button_20" at 720,420 size 80x60
   TextField "Text field_22" at 64,67 size 129x22
   AlarmView "Alarm view_1" at 60,90 size 680x320
   Button "Button_9" at 715,65 size 25x25
   TextField "Text field_37" at 360,54 size 120x25

screen "I0-State" 800x480
   TextField "Text field_3" at 325,5 size 300x40
   Button "Button_1" at 640,420 size 80x60
   Button "Button_4" at 160,420 size 80x60
   Button "HmiScreenItemData_3" at 400,420 size 80x60
   Button "Button_2" at 560,420 size 80x60
   Button "Button_6" at 720,420 size 80x60
   Button "HmiScreenItemData_2" at 240,420 size 80x60
   Button "HmiScreenItemData_4" at 320,420 size 80x60
   TextField "Text field_1" at 0,0 size 300x50
   DateTimeField "Date/time field_2" at 650,0 size 150x28
   DateTimeField "Date/time field_1" at 650,27 size 150x25
   Button "HmiScreenItemData_1" at 0,420 size 80x60
   Button "Button_3" at 480,420 size 80x60
   Button "Button_5" at 80,420 size 80x60
   Button "input_back" at 20,52 size 90x25
   Button "input_next" at 690,52 size 90x25
   Button "output_back" at 20,52 size 90x25
   Button "output_next" at 690,52 size 90x25
   TextField "Text field_2" at 20,85 size 330x22
   TextField "Text field_4" at 20,115 size 330x22
   TextField "Text field_5" at 20,145 size 330x22
   TextField "Text field_6" at 20,175 size 330x22
   TextField "Text field_7" at 20,205 size 330x22
   TextField "Text field_8" at 20,235 size 330x22
   TextField "Text field_9" at 20,265 size 330x22
   TextField "Text field_10" at 20,295 size 330x22
   TextField "Text field_11" at 20,325 size 330x22
   TextField "Text field_12" at 20,355 size 330x22
   TextField "Text field_13" at 20,385 size 330x22
   TextField "Text field_14" at 410,85 size 330x22
   TextField "Text field_15" at 410,115 size 330x22
   TextField "Text field_16" at 410,145 size 330x22
   TextField "Text field_17" at 410,175 size 330x22
   TextField "Text field_18" at 410,205 size 330x22
   TextField "Text field_19" at 410,235 size 330x22
   TextField "Text field_20" at 410,265 size 330x22
   TextField "Text field_21" at 410,295 size 330x22
   TextField "Text field_22" at 410,325 size 330x22
   TextField "Text field_23" at 410,355 size 330x22
   TextField "Text field_24" at 410,385 size 330x22
   Button "Button_11" at 0,420 size 80x60
   Button "Button_12" at 80,420 size 80x60
   Button "Button_13" at 160,420 size 80x60
   Button "Button_14" at 240,420 size 80x60
   Button "Button_15" at 320,420 size 80x60
   Button "Button_16" at 400,420 size 80x60
   Button "Button_17" at 480,420 size 80x60
   Button "Button_18" at 560,420 size 80x60
   Button "Button_19" at 640,420 size 80x60
   Button "Button_20" at 720,420 size 80x60
   TextField "Text field_25" at 64,67 size 129x22
   AlarmView "Alarm view_1" at 60,90 size 680x320
   Button "Button_9" at 715,65 size 25x25
   TextField "Text field_26" at 20,85 size 330x22
   TextField "Text field_27" at 20,115 size 330x22
   TextField "Text field_28" at 20,145 size 330x22
   TextField "Text field_29" at 20,175 size 330x22
   TextField "Text field_30" at 20,205 size 330x22
   TextField "Text field_31" at 20,235 size 330x22
   TextField "Text field_32" at 20,265 size 330x22
   TextField "Text field_33" at 20,295 size 330x22
   TextField "Text field_34" at 20,325 size 330x22
   TextField "Text field_48" at 21,85 size 330x22
   TextField "Text field_37" at 360,54 size 120x25

screen "Main_page" 800x480
   Button "HmiScreenItemData_1" at 80,420 size 80x60
   TextField "Text field_2" at 0,85 size 800x25
   TextField "Text field_3" at 325,5 size 300x40
   Button "Button_4" at 480,420 size 80x60
   Button "Button_5" at 640,420 size 80x60
   Button "Button_1" at 0,420 size 80x60
   Button "HmiScreenItemData_2" at 160,420 size 80x60
   Button "Button_2" at 400,420 size 80x60
   Button "Button_3" at 560,420 size 80x60
   Button "Button_6" at 720,420 size 80x60
   Button "HmiScreenItemData_3" at 240,420 size 80x60
   Button "HmiScreenItemData_4" at 320,420 size 80x60
   TextField "Text field_1" at 0,0 size 300x50
   DateTimeField "Date/time field_2" at 650,0 size 150x28
   DateTimeField "Date/time field_1" at 650,27 size 150x25
   SymbolicIOField "Symbolic I/O field_1" at 10,110 size 780x90
   Button "HmiScreenItemData_5" at 80,420 size 80x60
   GraphicView "Graphic view_1" at 320,228 size 180x180
   SymbolicIOField "Symbolic I/O field_6" at 169,51 size 169x32
   TextField "Text field_56" at 12,52 size 143x27
   Button "Button_21" at 720,420 size 80x60
   Button "Button_22" at 400,420 size 80x60
   Button "Button_11" at 0,420 size 80x60
   Button "Button_13" at 160,420 size 80x60
   Button "Button_14" at 240,420 size 80x60
   Button "Button_15" at 320,420 size 80x60
   Button "Button_16" at 400,420 size 80x60
   Button "Button_17" at 480,420 size 80x60
   Button "Button_18" at 560,420 size 80x60
   Button "Button_19" at 640,420 size 80x60
   Button "Button_20" at 720,420 size 80x60
   Button "Button_12" at 80,420 size 80x60
   TextField "Text field_5" at 64,67 size 129x22
   AlarmView "Alarm view_1" at 60,90 size 680x320
   Button "Button_9" at 715,65 size 25x25
   SymbolicIOField "Symbolic I/O field_2" at 0,170 size 800x110
   SymbolicIOField "Symbolic I/O field_3" at 0,170 size 800x110
   SymbolicIOField "Symbolic I/O field_4" at 0,170 size 800x110
   SymbolicIOField "Symbolic I/O field_5" at 0,170 size 800x110
   Button "Button_7" at 486,333 size 130x50
   Button "Button_10" at 213,333 size 130x50
   Button "Button_8" at 350,333 size 130x50
   TextField "Text field_37" at 360,54 size 120x25
   TextField "Text field_4" at 302,290 size 237x43

screen "Scanner" 800x480
   TextField "Text field_3" at 325,5 size 300x40
   IOField "I/O field_1" at 10,120 size 780x32
   TextField "Text field_2" at 10,88 size 141x22
   Button "Button_1" at 640,420 size 80x60
   Button "HmiScreenItemData_3" at 400,420 size 80x60
   Button "Button_2" at 560,420 size 80x60
   Button "Button_6" at 720,420 size 80x60
   DateTimeField "Date/time field_2" at 650,0 size 150x28
   TextField "Text field_1" at 0,0 size 300x50
   DateTimeField "Date/time field_1" at 650,27 size 150x25
   Button "HmiScreenItemData_2" at 240,420 size 80x60
   Button "HmiScreenItemData_4" at 320,420 size 80x60
   Button "HmiScreenItemData_1" at 0,420 size 80x60
   Button "HmiScreenItemData_5" at 480,420 size 80x60
   Button "HmiScreenItemData_6" at 160,420 size 80x60
   Button "HmiScreenItemData_7" at 80,420 size 80x60
   Button "Button_3" at 10,165 size 96x32
   Button "Button_11" at 0,420 size 80x60
   Button "Button_12" at 80,420 size 80x60
   Button "Button_13" at 160,420 size 80x60
   Button "Button_14" at 240,420 size 80x60
   Button "Button_15" at 320,420 size 80x60
   Button "Button_16" at 400,420 size 80x60
   Button "Button_17" at 480,420 size 80x60
   Button "Button_18" at 560,420 size 80x60
   Button "Button_19" at 640,420 size 80x60
   Button "Button_20" at 720,420 size 80x60
   TextField "Text field_5" at 64,67 size 129x22
   AlarmView "Alarm view_1" at 60,90 size 680x320
   Button "Button_9" at 715,65 size 25x25
   TextField "Text field_37" at 360,54 size 120x25

screen "Manual" 800x480
   TextField "Text field_3" at 325,5 size 300x40
   Button "Button_12" at 730,85 size 50x50
   Button "Button_1" at 640,420 size 80x60
   Button "HmiScreenItemData_1" at 0,420 size 80x60
   Button "Button_2" at 560,420 size 80x60
   Button "Button_6" at 720,420 size 80x60
   Button "Button_34" at 400,420 size 80x60
   Button "HmiScreenItemData_3" at 240,420 size 80x60
   Button "HmiScreenItemData_4" at 320,420 size 80x60
   DateTimeField "Date/time field_2" at 650,0 size 150x28
   DateTimeField "Date/time field_1" at 650,27 size 150x25
   Button "Button_5" at 160,420 size 80x60
   Button "Button_3" at 480,420 size 80x60
   Button "Button_7" at 80,420 size 80x60
   Button "Button_4" at 21,85 size 50x50
   TextField "Text field_1" at 0,0 size 300x50
   Button "Button_23" at 0,420 size 80x60
   Button "Button_24" at 80,420 size 80x60
   Button "Button_25" at 160,420 size 80x60
   Button "Button_26" at 240,420 size 80x60
   Button "Button_27" at 320,420 size 80x60
   Button "Button_28" at 400,420 size 80x60
   Button "Button_29" at 480,420 size 80x60
   Button "Button_30" at 560,420 size 80x60
   Button "Button_31" at 640,420 size 80x60
   Button "Button_32" at 720,420 size 80x60
   AlarmView "Alarm view_1" at 60,90 size 680x320
   TextField "Text field_8" at 64,67 size 129x22
   Button "Button_33" at 715,65 size 25x25
   Switch "Switch_1" at 717,149 size 64x32
   Switch "Switch_2" at 717,185 size 64x32
   TextField "Text field_7" at 493,149 size 200x32
   TextField "Text field_9" at 493,181 size 200x32
   Switch "Switch_8" at 300,149 size 64x32
   Switch "Switch_9" at 300,185 size 64x32
   Switch "Switch_10" at 300,221 size 64x32
   Switch "Switch_11" at 300,257 size 64x32
   Switch "Switch_12" at 300,293 size 64x32
   Switch "Switch_13" at 301,328 size 64x32
   Switch "Switch_14" at 302,364 size 64x32
   TextField "Text field_15" at 76,149 size 200x32
   TextField "Text field_16" at 76,181 size 200x32
   TextField "Text field_17" at 75,221 size 200x32
   TextField "Text field_18" at 37,289 size 239x32
   TextField "Text field_19" at 26,257 size 250x32
   TextField "Text field_20" at 29,328 size 247x32
   TextField "Text field_21" at 44,360 size 232x32
   TextField "Text field_37" at 360,54 size 120x25

screen "System" 800x480
   TextField "Text field_3" at 325,5 size 300x40
   TextField "Text field_2" at 300,85 size 200x27
   Button "Button_4" at 10,290 size 170x60
   Button "Button_5" at 10,355 size 170x60
   Button "Button_7" at 213,290 size 170x60
   Button "Button_8" at 416,290 size 170x60
   Button "Button_9" at 620,290 size 170x60
   Button "Button_11" at 213,355 size 170x60
   Button "Button_12" at 416,355 size 170x60
   Button "Button_13" at 620,355 size 170x60
   AlarmView "Alarm view_1" at 10,116 size 780x169
   Button "HmiScreenItemData_1" at 0,420 size 80x60
   Button "Button_3" at 160,420 size 80x60
   Button "Button_14" at 240,420 size 80x60
   Button "Button_15" at 320,420 size 80x60
   Button "Button_16" at 400,420 size 80x60
   Button "Button_2" at 560,420 size 80x60
   Button "Button_1" at 640,420 size 80x60
   Button "Button_6" at 720,420 size 80x60
   TextField "Text field_1" at 0,0 size 300x50
   DateTimeField "Date/time field_2" at 650,0 size 150x28
   DateTimeField "Date/time field_1" at 650,27 size 150x25
   Button "Button_10" at 80,420 size 80x60
   Button "Button_17" at 480,420 size 80x60
   TextField "Text field_37" at 360,54 size 120x25

screen "type" 800x480
   TextField "Text field_3" at 325,5 size 300x40
   Button "Button_1" at 640,420 size 80x60
   Button "HmiScreenItemData_1" at 0,420 size 80x60
   Button "Button_6" at 720,420 size 80x60
   Button "Button_34" at 400,420 size 80x60
   Button "HmiScreenItemData_4" at 320,420 size 80x60
   TextField "Text field_1" at 0,0 size 300x50
   DateTimeField "Date/time field_2" at 650,0 size 150x28
   DateTimeField "Date/time field_1" at 650,27 size 150x25
   Button "Button_5" at 160,420 size 80x60
   Button "Button_3" at 480,420 size 80x60
   Button "Button_7" at 80,420 size 80x60
   Button "Button_2" at 560,420 size 80x60
   SymbolicIOField "Symbolic I/O field_1" at 33,194 size 310x65
   TextField "Text field_2" at 33,159 size 192x27
   Button "Button_4" at 355,195 size 90x65
   SymbolicIOField "Symbolic I/O field_2" at 457,195 size 310x65
   TextField "Text field_4" at 457,159 size 225x27
   Button "HmiScreenItemData_2" at 240,420 size 80x60
   TextField "Text field_37" at 360,54 size 120x25
*)

(* ===== HMI "HMI_RT_5" =====
connection "HMI_Connection_5": ETHERNET, SMART_S7_1500_OMS
